(* Logix 5000 project; controller FV vendor 1 type 14 code 217 rev 31.11; software revision 31.00; part 31 of 63 *)
(* tags used below, declared in another part *)
   CWD : CHECKWORD_FLAGS;
   FR_BEACON1 : PlantItem;   // BEACON1
   FR_data_file_value_to_move : DINT;
   FR_F202 : REAL[20];
   FR_F203 : REAL[40];
   FR_N120 : INT[265];   // YEAST CROP Yeast Cropping Main
   FR_N14 : INT[265];   // MVFV CIP Comms to MVFV CIP Un it PLC
   FR_N140 : INT[265];   // CIP
   FR_N160 : INT[265];   // VESSEL Vessel Working Direc tory
   FR_N20 : INT[265];   // GENERAL General Purpose Setp oints
   FR_N30 : INT[265];   // FV30
   FR_N7 : INT[265];   // INTEGER
   FR_N99 : INT[265];   // COMMENT Comment Lines
   FR_T121 : TIMER[255];   // YEAST CROP
   scale_analog_result : REAL;
(* FR_Common, continued *)

ROUTINE FR_VESSEL_160   (* ladder *)
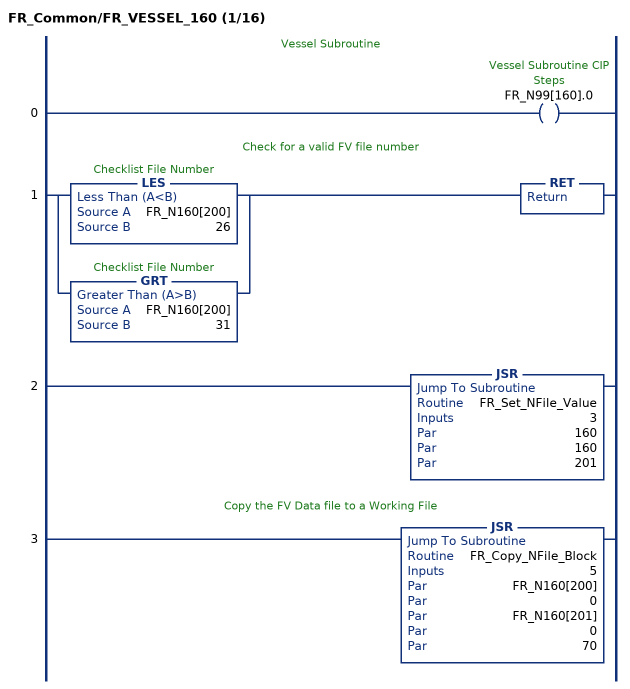
   // Vessel Subroutine
   0: OTE(FR_N99[160].0);
   // Check for a valid FV file number
   1: [LES(FR_N160[200],26) ,GRT(FR_N160[200],31) ]RET();
   2: JSR(FR_Set_NFile_Value,3,160,160,201);
   // Copy the FV Data file to a Working File
   3: JSR(FR_Copy_NFile_Block,5,FR_N160[200],0,FR_N160[201],0,70);
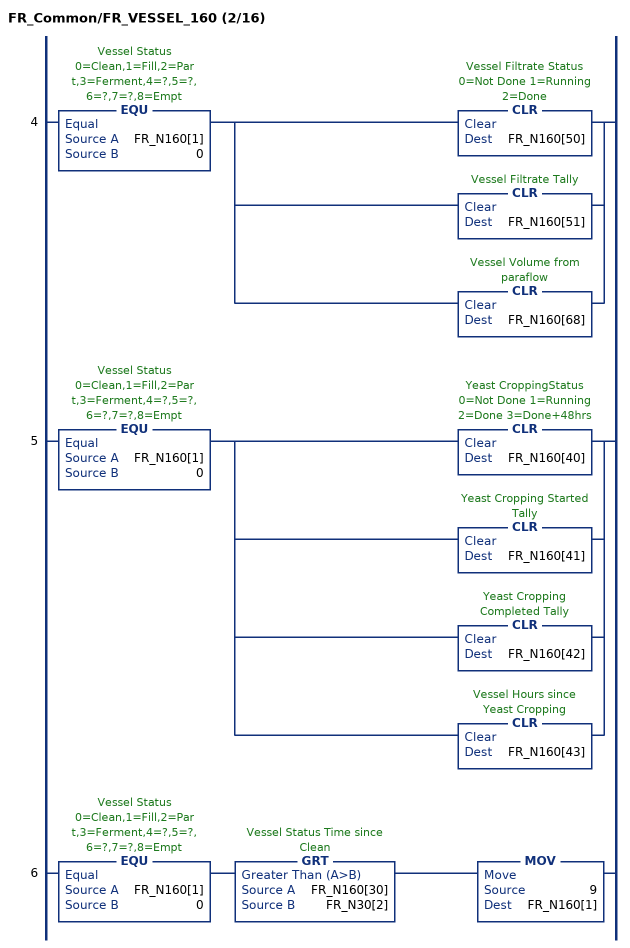
   4: EQU(FR_N160[1],0)[CLR(FR_N160[50]) ,CLR(FR_N160[51]) ,CLR(FR_N160[68]) ];
   5: EQU(FR_N160[1],0)[CLR(FR_N160[40]) ,CLR(FR_N160[41]) ,CLR(FR_N160[42]) ,CLR(FR_N160[43]) ];
   6: EQU(FR_N160[1],0)GRT(FR_N160[30],FR_N30[2])MOV(9,FR_N160[1]);
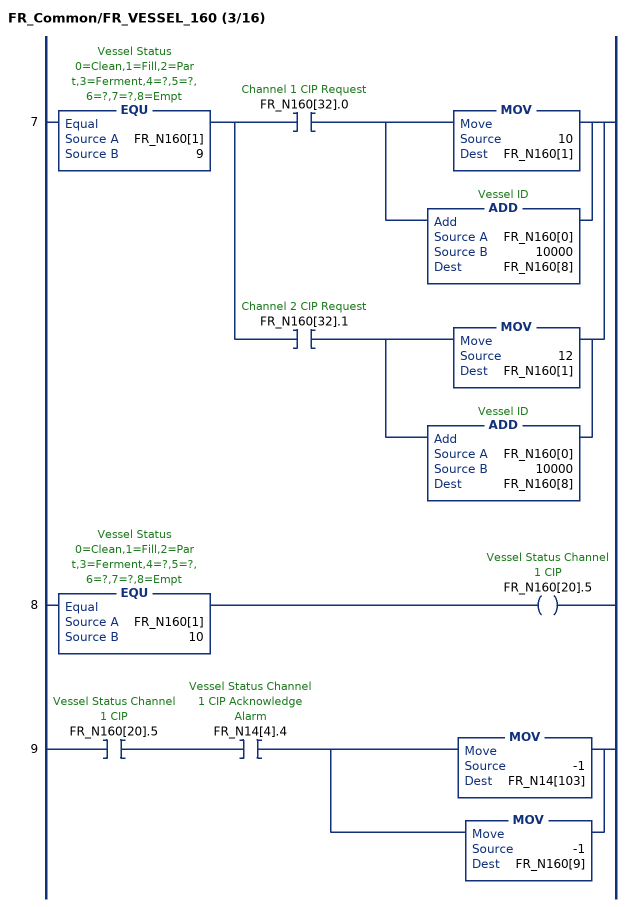
   7: EQU(FR_N160[1],9)[XIC(FR_N160[32].0) [MOV(10,FR_N160[1]) ,ADD(FR_N160[0],10000,FR_N160[8]) ] ,XIC(FR_N160[32].1) [MOV(12,FR_N160[1]) ,ADD(FR_N160[0],10000,FR_N160[8]) ] ];
   8: EQU(FR_N160[1],10)OTE(FR_N160[20].5);
   9: XIC(FR_N160[20].5)XIC(FR_N14[4].4)[MOV(-1,FR_N14[103]) ,MOV(-1,FR_N160[9]) ];
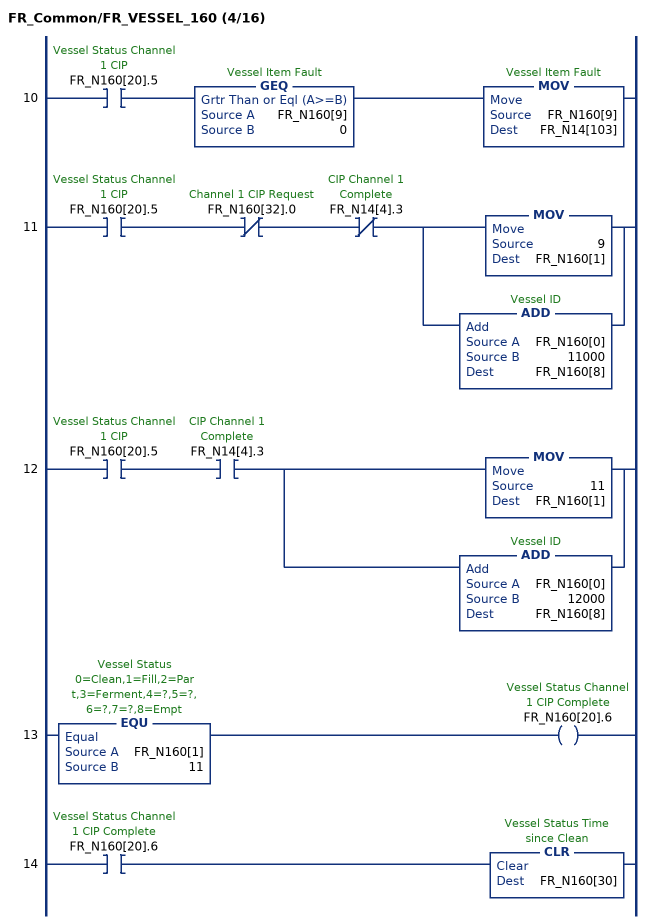
   10: XIC(FR_N160[20].5)GEQ(FR_N160[9],0)MOV(FR_N160[9],FR_N14[103]);
   11: XIC(FR_N160[20].5)XIO(FR_N160[32].0)XIO(FR_N14[4].3)[MOV(9,FR_N160[1]) ,ADD(FR_N160[0],11000,FR_N160[8]) ];
   12: XIC(FR_N160[20].5)XIC(FR_N14[4].3)[MOV(11,FR_N160[1]) ,ADD(FR_N160[0],12000,FR_N160[8]) ];
   13: EQU(FR_N160[1],11)OTE(FR_N160[20].6);
   14: XIC(FR_N160[20].6)CLR(FR_N160[30]);
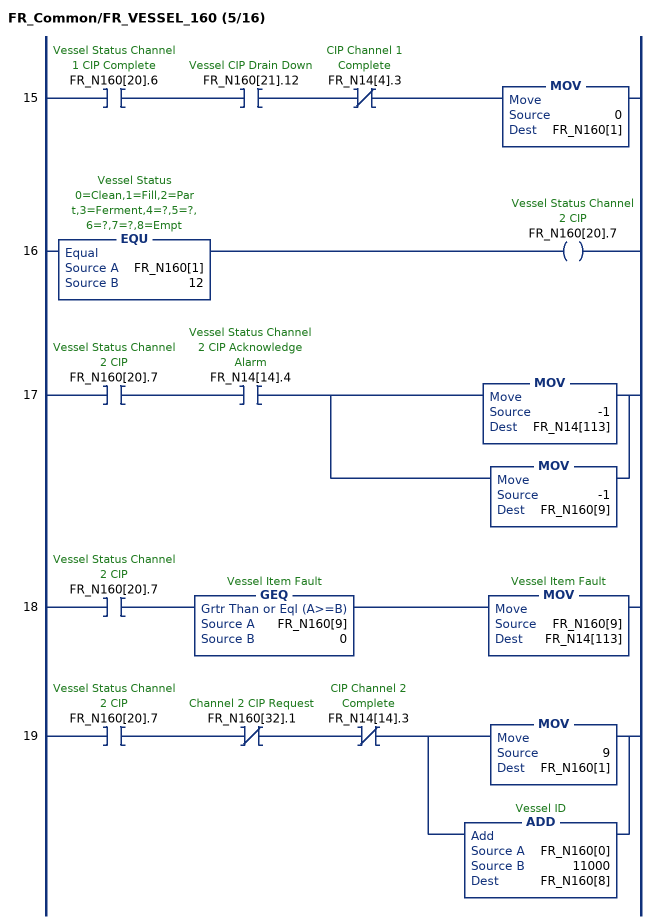
   15: XIC(FR_N160[20].6)XIC(FR_N160[21].12)XIO(FR_N14[4].3)MOV(0,FR_N160[1]);
   16: EQU(FR_N160[1],12)OTE(FR_N160[20].7);
   17: XIC(FR_N160[20].7)XIC(FR_N14[14].4)[MOV(-1,FR_N14[113]) ,MOV(-1,FR_N160[9]) ];
   18: XIC(FR_N160[20].7)GEQ(FR_N160[9],0)MOV(FR_N160[9],FR_N14[113]);
   19: XIC(FR_N160[20].7)XIO(FR_N160[32].1)XIO(FR_N14[14].3)[MOV(9,FR_N160[1]) ,ADD(FR_N160[0],11000,FR_N160[8]) ];
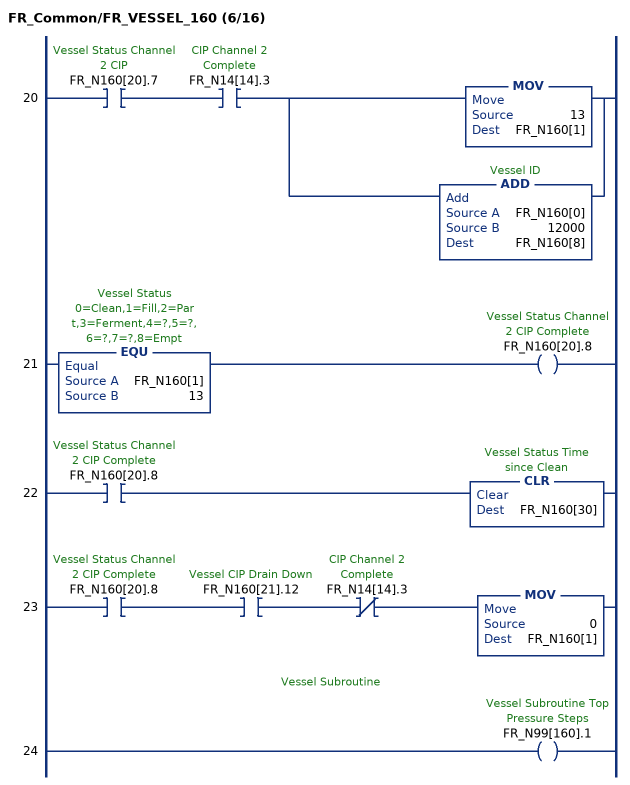
   20: XIC(FR_N160[20].7)XIC(FR_N14[14].3)[MOV(13,FR_N160[1]) ,ADD(FR_N160[0],12000,FR_N160[8]) ];
   21: EQU(FR_N160[1],13)OTE(FR_N160[20].8);
   22: XIC(FR_N160[20].8)CLR(FR_N160[30]);
   23: XIC(FR_N160[20].8)XIC(FR_N160[21].12)XIO(FR_N14[14].3)MOV(0,FR_N160[1]);
   // Vessel Subroutine
   24: OTE(FR_N99[160].1);
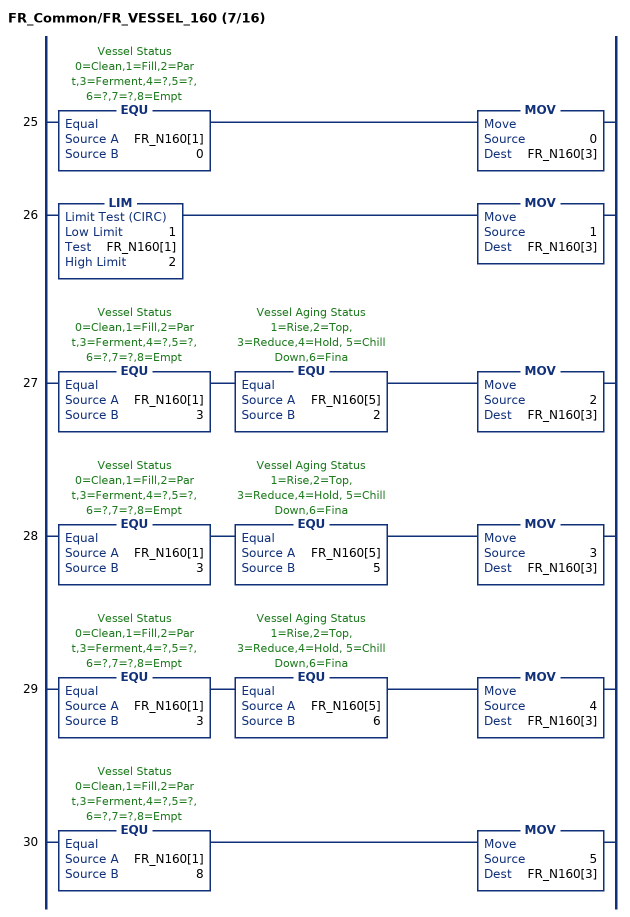
   25: EQU(FR_N160[1],0)MOV(0,FR_N160[3]);
   26: LIM(1,FR_N160[1],2)MOV(1,FR_N160[3]);
   27: EQU(FR_N160[1],3)EQU(FR_N160[5],2)MOV(2,FR_N160[3]);
   28: EQU(FR_N160[1],3)EQU(FR_N160[5],5)MOV(3,FR_N160[3]);
   29: EQU(FR_N160[1],3)EQU(FR_N160[5],6)MOV(4,FR_N160[3]);
   30: EQU(FR_N160[1],8)MOV(5,FR_N160[3]);
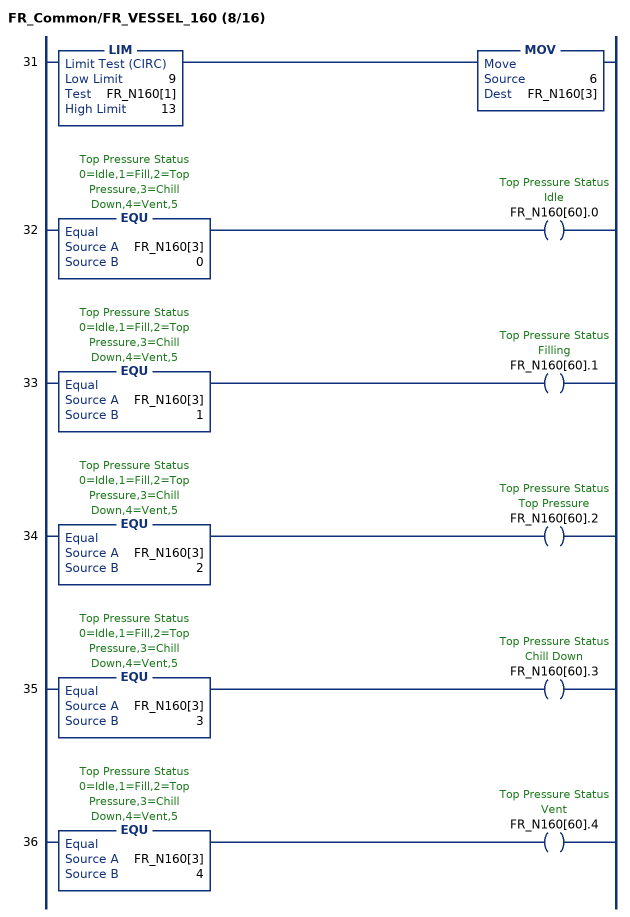
   31: LIM(9,FR_N160[1],13)MOV(6,FR_N160[3]);
   32: EQU(FR_N160[3],0)OTE(FR_N160[60].0);
   33: EQU(FR_N160[3],1)OTE(FR_N160[60].1);
   34: EQU(FR_N160[3],2)OTE(FR_N160[60].2);
   35: EQU(FR_N160[3],3)OTE(FR_N160[60].3);
   36: EQU(FR_N160[3],4)OTE(FR_N160[60].4);
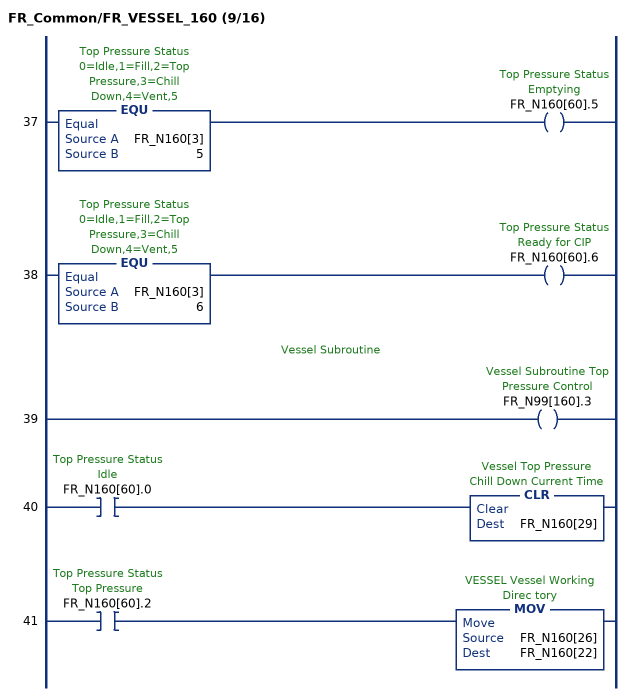
   37: EQU(FR_N160[3],5)OTE(FR_N160[60].5);
   38: EQU(FR_N160[3],6)OTE(FR_N160[60].6);
   // Vessel Subroutine
   39: OTE(FR_N99[160].3);
   40: XIC(FR_N160[60].0)CLR(FR_N160[29]);
   41: XIC(FR_N160[60].2)MOV(FR_N160[26],FR_N160[22]);
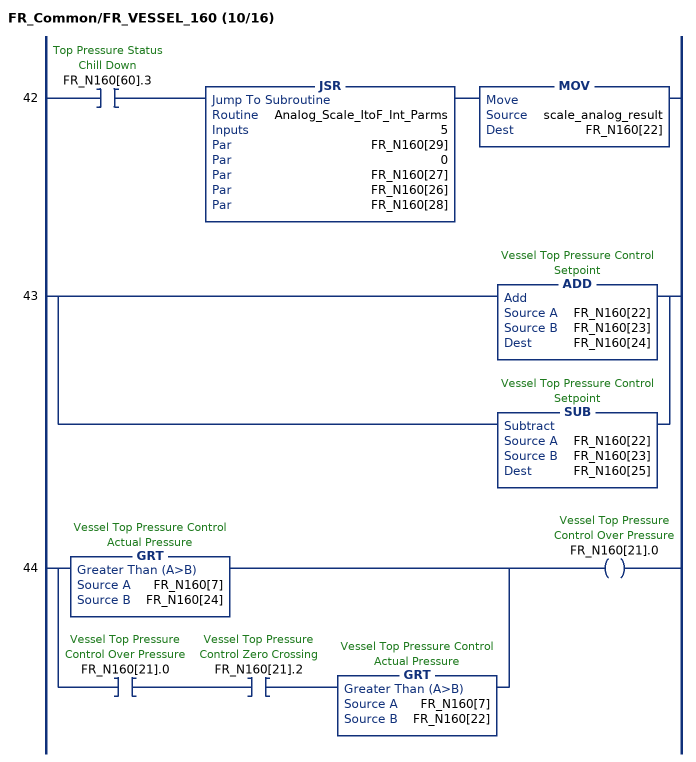
   42: XIC(FR_N160[60].3)JSR(Analog_Scale_ItoF_Int_Parms,5,FR_N160[29],0,FR_N160[27],FR_N160[26],FR_N160[28])MOV(scale_analog_result,FR_N160[22]);
   43: [ADD(FR_N160[22],FR_N160[23],FR_N160[24]) ,SUB(FR_N160[22],FR_N160[23],FR_N160[25]) ];
   44: [GRT(FR_N160[7],FR_N160[24]) ,XIC(FR_N160[21].0) XIC(FR_N160[21].2) GRT(FR_N160[7],FR_N160[22]) ]OTE(FR_N160[21].0);
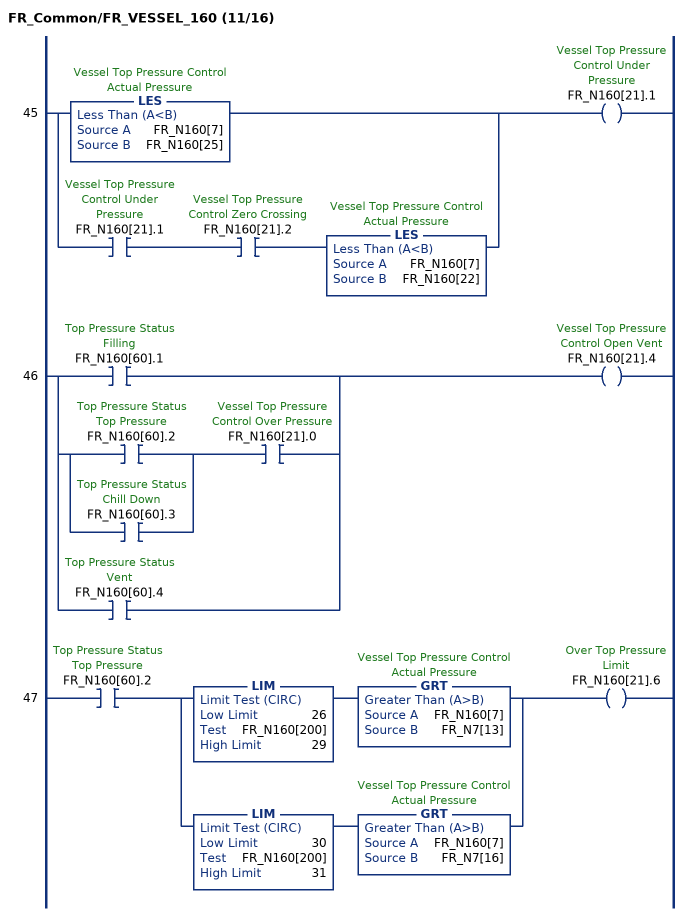
   45: [LES(FR_N160[7],FR_N160[25]) ,XIC(FR_N160[21].1) XIC(FR_N160[21].2) LES(FR_N160[7],FR_N160[22]) ]OTE(FR_N160[21].1);
   46: [XIC(FR_N160[60].1) ,[XIC(FR_N160[60].2) ,XIC(FR_N160[60].3) ] XIC(FR_N160[21].0) ,XIC(FR_N160[60].4) ]OTE(FR_N160[21].4);
   47: XIC(FR_N160[60].2)[LIM(26,FR_N160[200],29) GRT(FR_N160[7],FR_N7[13]) ,LIM(30,FR_N160[200],31) GRT(FR_N160[7],FR_N7[16]) ]OTE(FR_N160[21].6);
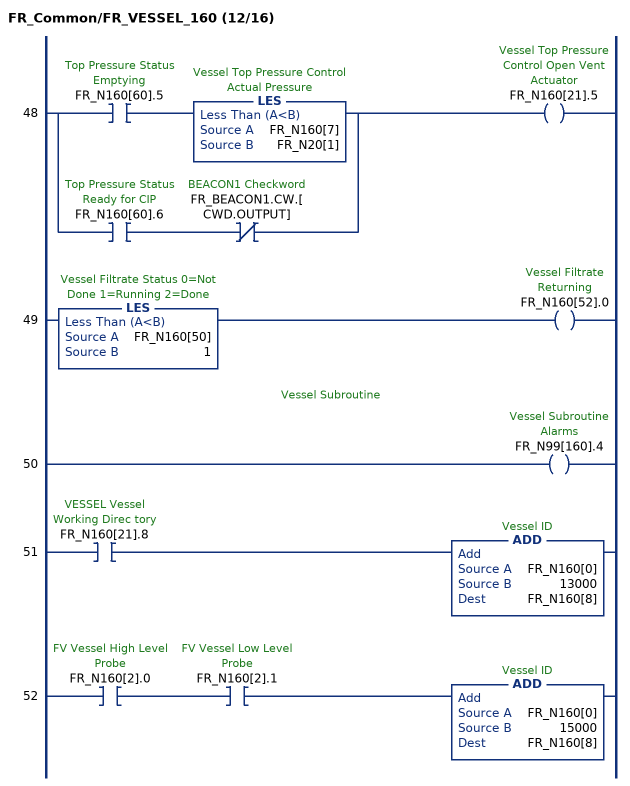
   48: [XIC(FR_N160[60].5) LES(FR_N160[7],FR_N20[1]) ,XIC(FR_N160[60].6) XIO(FR_BEACON1.CW.[CWD.OUTPUT]) ]OTE(FR_N160[21].5);
   49: LES(FR_N160[50],1)OTE(FR_N160[52].0);
   // Vessel Subroutine
   50: OTE(FR_N99[160].4);
   51: XIC(FR_N160[21].8)ADD(FR_N160[0],13000,FR_N160[8]);
   52: XIC(FR_N160[2].0)XIC(FR_N160[2].1)ADD(FR_N160[0],15000,FR_N160[8]);
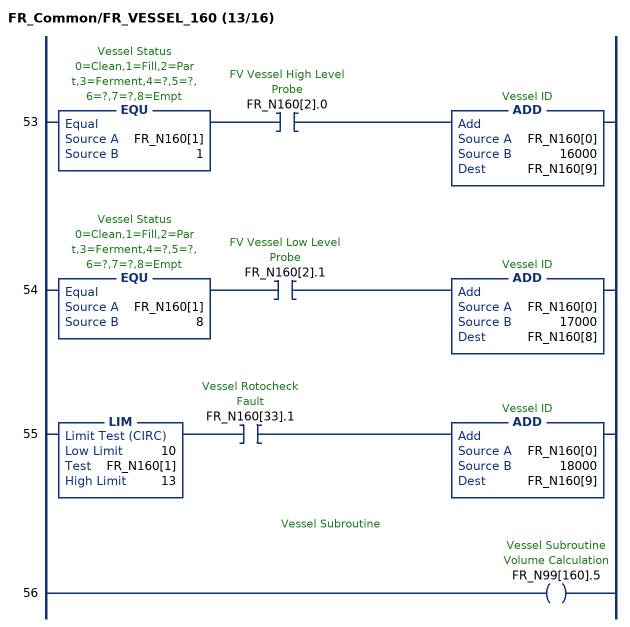
   53: EQU(FR_N160[1],1)XIC(FR_N160[2].0)ADD(FR_N160[0],16000,FR_N160[9]);
   54: EQU(FR_N160[1],8)XIC(FR_N160[2].1)ADD(FR_N160[0],17000,FR_N160[8]);
   55: LIM(10,FR_N160[1],13)XIC(FR_N160[33].1)ADD(FR_N160[0],18000,FR_N160[9]);
   // Vessel Subroutine
   56: OTE(FR_N99[160].5);
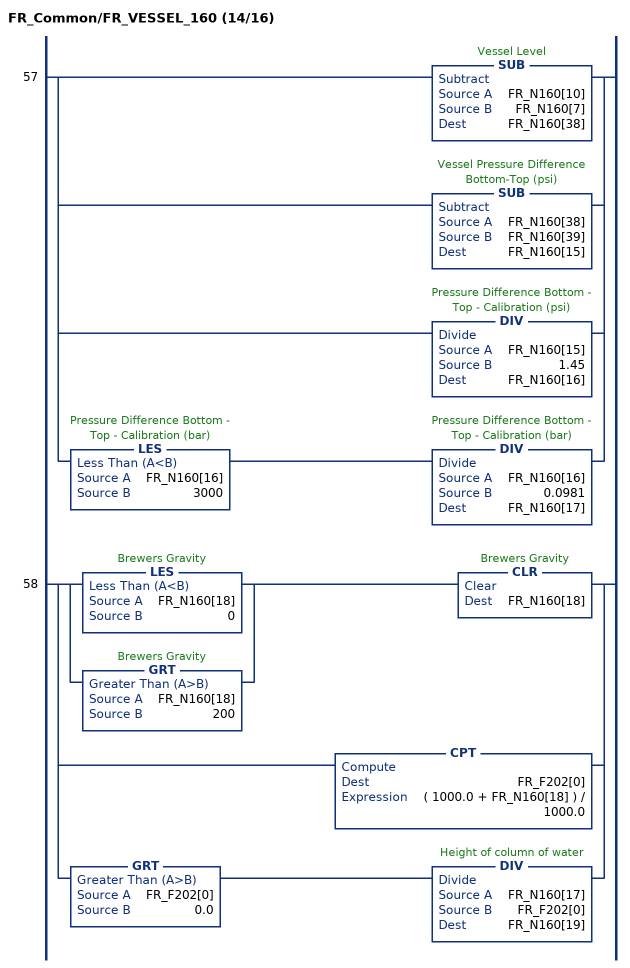
   57: [SUB(FR_N160[10],FR_N160[7],FR_N160[38]) ,SUB(FR_N160[38],FR_N160[39],FR_N160[15]) ,DIV(FR_N160[15],1.45,FR_N160[16]) ,LES(FR_N160[16],3000) DIV(FR_N160[16],0.0981,FR_N160[17]) ];
   58: [[LES(FR_N160[18],0) ,GRT(FR_N160[18],200) ] CLR(FR_N160[18]) ,CPT(FR_F202[0],( 1000.0 + FR_N160[18] ) / 1000.0) ,GRT(FR_F202[0],0.0) DIV(FR_N160[17],FR_F202[0],FR_N160[19]) ];
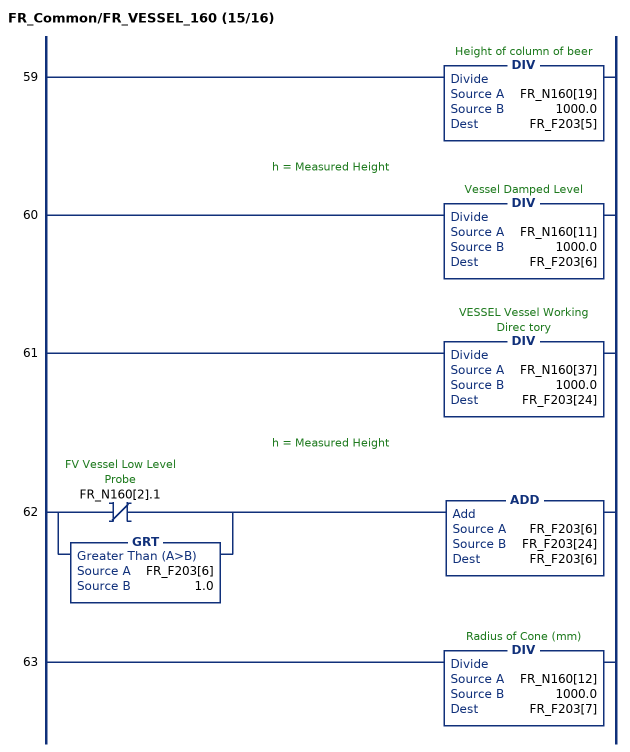
   59: DIV(FR_N160[19],1000.0,FR_F203[5]);
   // h = Measured Height
   60: DIV(FR_N160[11],1000.0,FR_F203[6]);
   61: DIV(FR_N160[37],1000.0,FR_F203[24]);
   // h = Measured Height
   62: [XIO(FR_N160[2].1) ,GRT(FR_F203[6],1.0) ]ADD(FR_F203[6],FR_F203[24],FR_F203[6]);
   63: DIV(FR_N160[12],1000.0,FR_F203[7]);
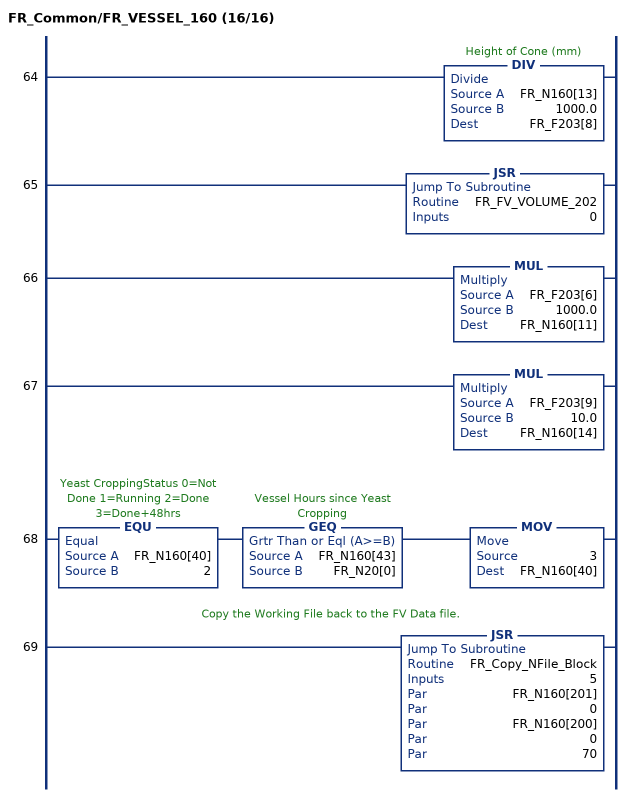
   64: DIV(FR_N160[13],1000.0,FR_F203[8]);
   65: JSR(FR_FV_VOLUME_202,0);
   66: MUL(FR_F203[6],1000.0,FR_N160[11]);
   67: MUL(FR_F203[9],10.0,FR_N160[14]);
   68: EQU(FR_N160[40],2)GEQ(FR_N160[43],FR_N20[0])MOV(3,FR_N160[40]);
   // Copy the Working File back to the FV Data file.
   69: JSR(FR_Copy_NFile_Block,5,FR_N160[201],0,FR_N160[200],0,70);
END_ROUTINE

ROUTINE FR_YEAST_121   (* ladder *)
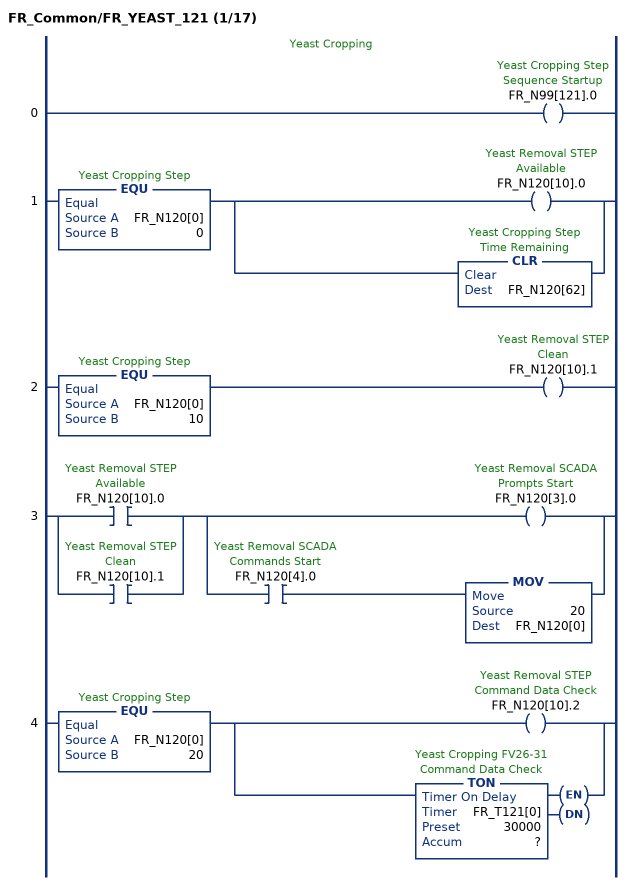
   // Yeast Cropping
   0: OTE(FR_N99[121].0);
   1: EQU(FR_N120[0],0)[OTE(FR_N120[10].0) ,CLR(FR_N120[62]) ];
   2: EQU(FR_N120[0],10)OTE(FR_N120[10].1);
   3: [XIC(FR_N120[10].0) ,XIC(FR_N120[10].1) ][OTE(FR_N120[3].0) ,XIC(FR_N120[4].0) MOV(20,FR_N120[0]) ];
   4: EQU(FR_N120[0],20)[OTE(FR_N120[10].2) ,TON(FR_T121[0],?,?) ];
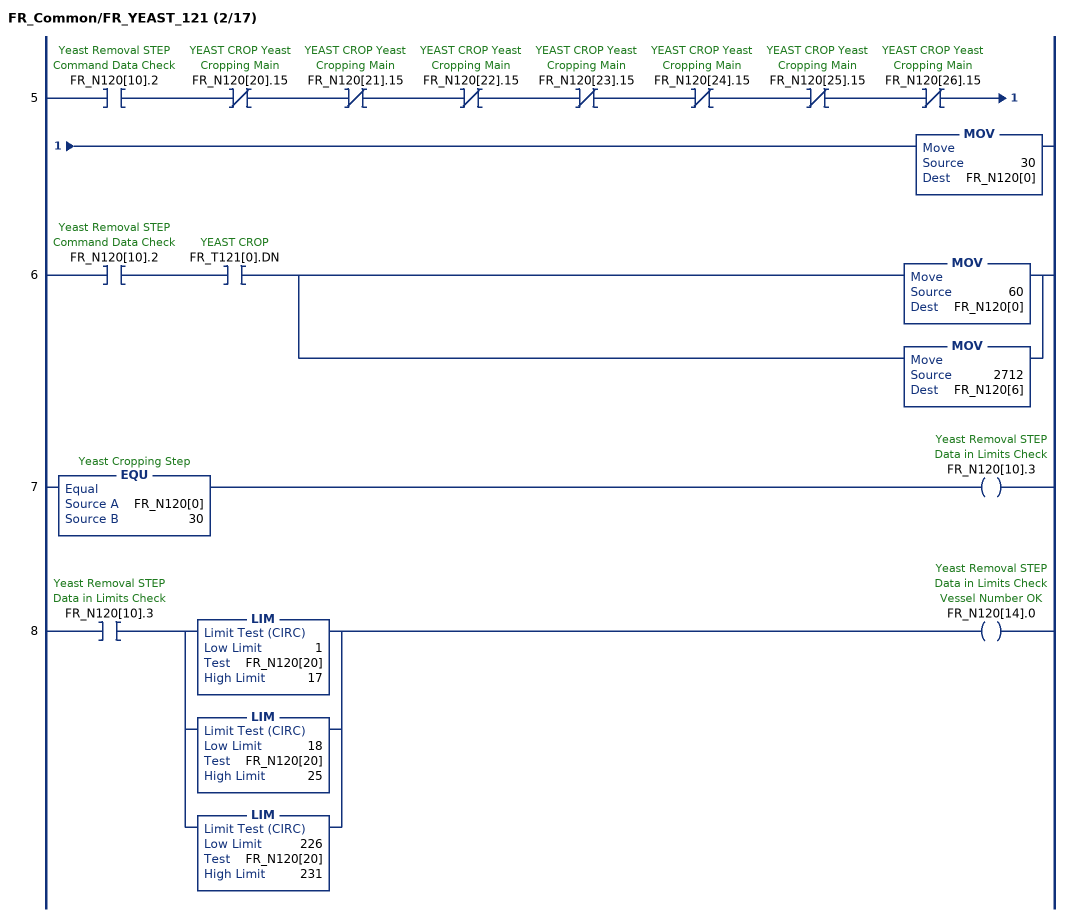
   5: XIC(FR_N120[10].2)XIO(FR_N120[20].15)XIO(FR_N120[21].15)XIO(FR_N120[22].15)XIO(FR_N120[23].15)XIO(FR_N120[24].15)XIO(FR_N120[25].15)XIO(FR_N120[26].15)MOV(30,FR_N120[0]);
   6: XIC(FR_N120[10].2)XIC(FR_T121[0].DN)[MOV(60,FR_N120[0]) ,MOV(2712,FR_N120[6]) ];
   7: EQU(FR_N120[0],30)OTE(FR_N120[10].3);
   8: XIC(FR_N120[10].3)[LIM(1,FR_N120[20],17) ,LIM(18,FR_N120[20],25) ,LIM(226,FR_N120[20],231) ]OTE(FR_N120[14].0);
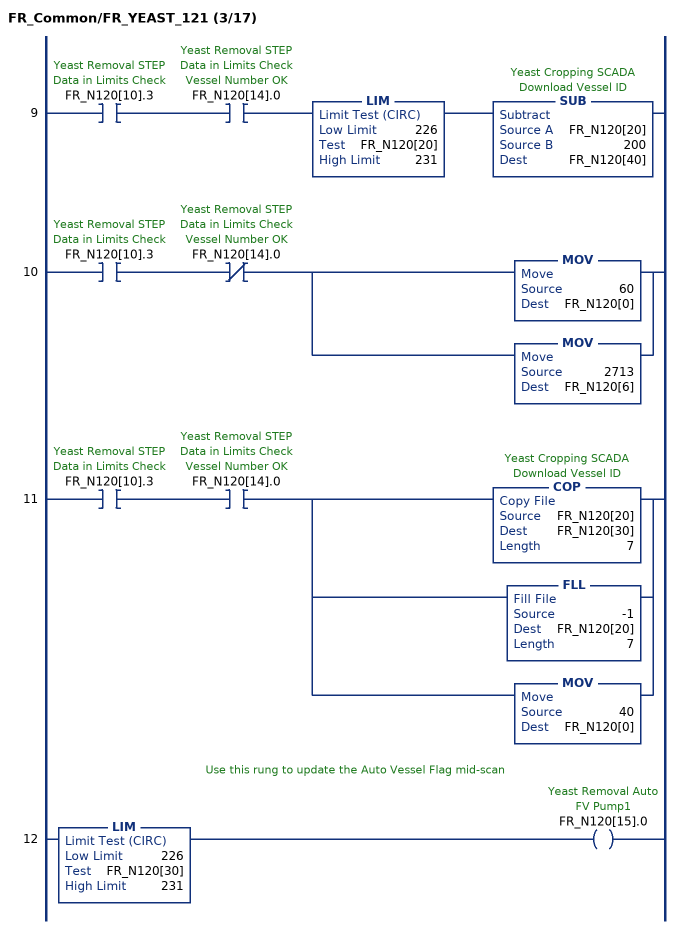
   9: XIC(FR_N120[10].3)XIC(FR_N120[14].0)LIM(226,FR_N120[20],231)SUB(FR_N120[20],200,FR_N120[40]);
   10: XIC(FR_N120[10].3)XIO(FR_N120[14].0)[MOV(60,FR_N120[0]) ,MOV(2713,FR_N120[6]) ];
   11: XIC(FR_N120[10].3)XIC(FR_N120[14].0)[COP(FR_N120[20],FR_N120[30],7) ,FLL(-1,FR_N120[20],7) ,MOV(40,FR_N120[0]) ];
   // Use this rung to update the Auto Vessel Flag mid-scan
   12: LIM(226,FR_N120[30],231)OTE(FR_N120[15].0);
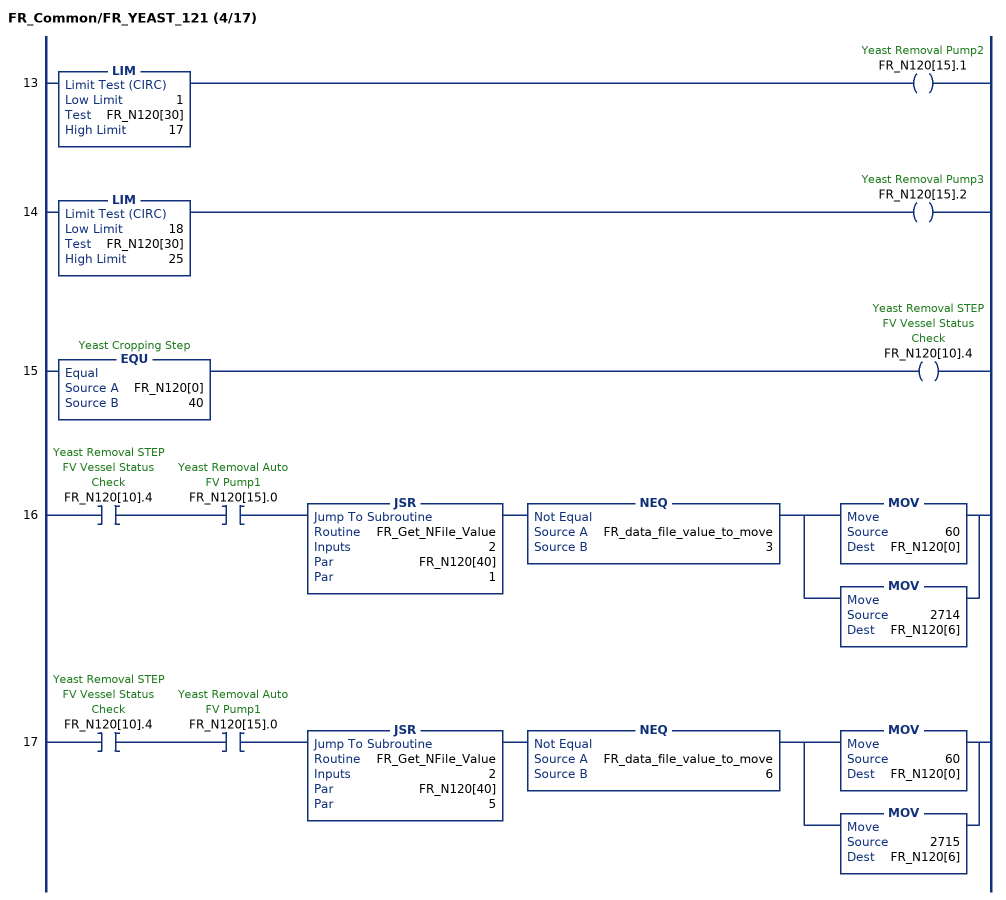
   13: LIM(1,FR_N120[30],17)OTE(FR_N120[15].1);
   14: LIM(18,FR_N120[30],25)OTE(FR_N120[15].2);
   15: EQU(FR_N120[0],40)OTE(FR_N120[10].4);
   16: XIC(FR_N120[10].4)XIC(FR_N120[15].0)JSR(FR_Get_NFile_Value,2,FR_N120[40],1)NEQ(FR_data_file_value_to_move,3)[MOV(60,FR_N120[0]) ,MOV(2714,FR_N120[6]) ];
   17: XIC(FR_N120[10].4)XIC(FR_N120[15].0)JSR(FR_Get_NFile_Value,2,FR_N120[40],5)NEQ(FR_data_file_value_to_move,6)[MOV(60,FR_N120[0]) ,MOV(2715,FR_N120[6]) ];
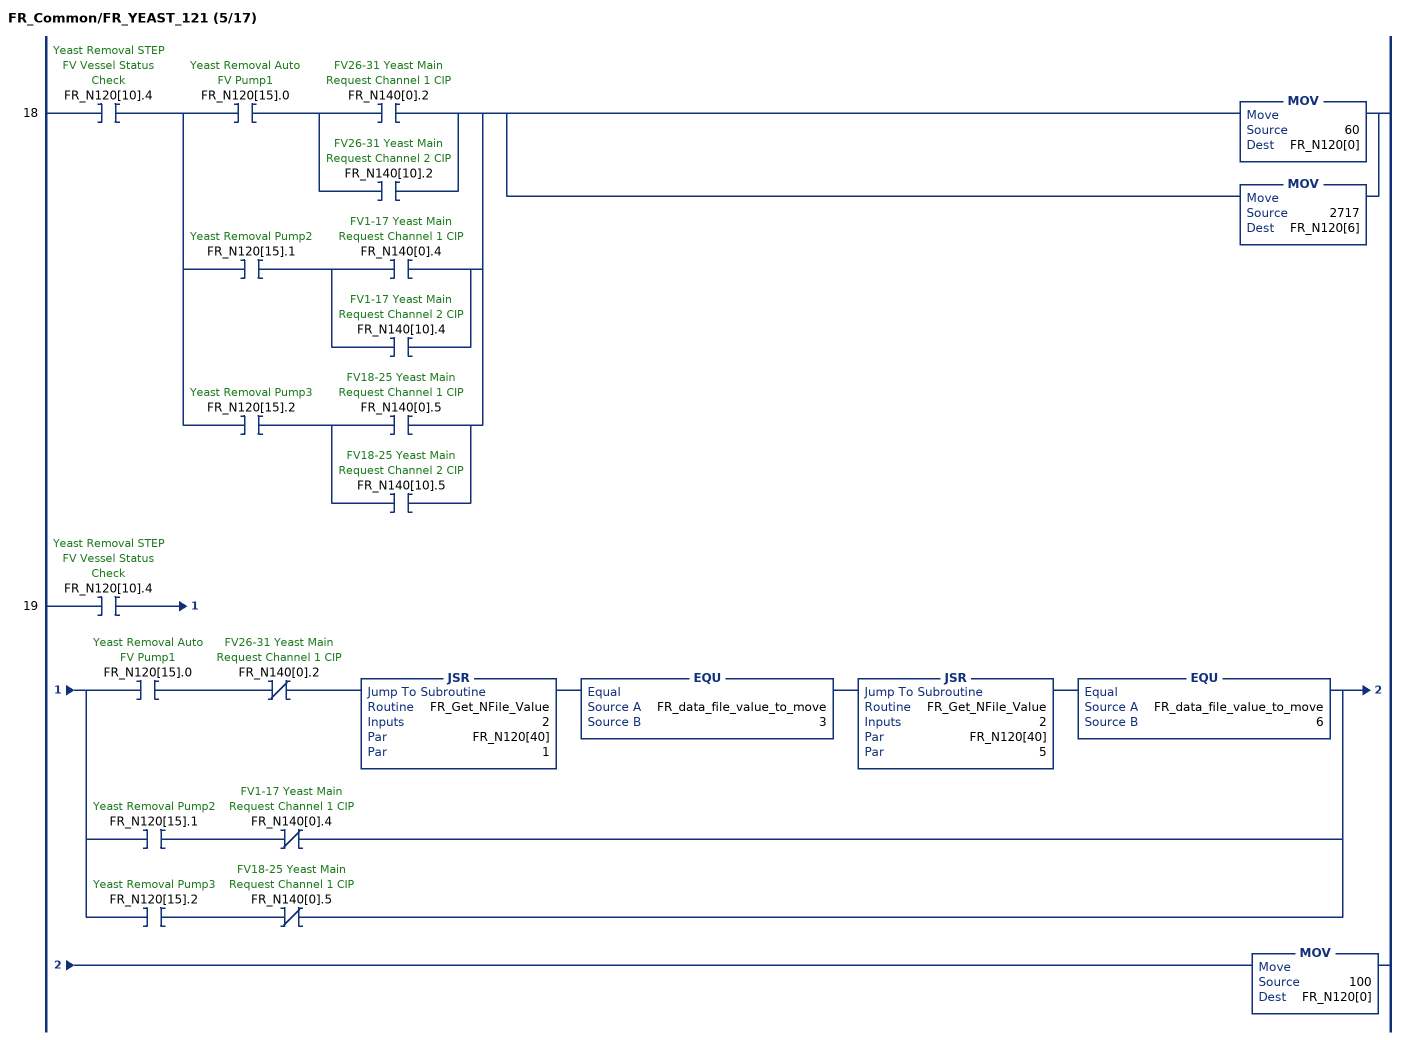
   18: XIC(FR_N120[10].4)[XIC(FR_N120[15].0) [XIC(FR_N140[0].2) ,XIC(FR_N140[10].2) ] ,XIC(FR_N120[15].1) [XIC(FR_N140[0].4) ,XIC(FR_N140[10].4) ] ,XIC(FR_N120[15].2) [XIC(FR_N140[0].5) ,XIC(FR_N140[10].5) ] ][MOV(60,FR_N120[0]) ,MOV(2717,FR_N120[6]) ];
   19: XIC(FR_N120[10].4)[XIC(FR_N120[15].0) XIO(FR_N140[0].2) JSR(FR_Get_NFile_Value,2,FR_N120[40],1) EQU(FR_data_file_value_to_move,3) JSR(FR_Get_NFile_Value,2,FR_N120[40],5) EQU(FR_data_file_value_to_move,6) ,XIC(FR_N120[15].1) XIO(FR_N140[0].4) ,XIC(FR_N120[15].2) XIO(FR_N140[0].5) ]MOV(100,FR_N120[0]);
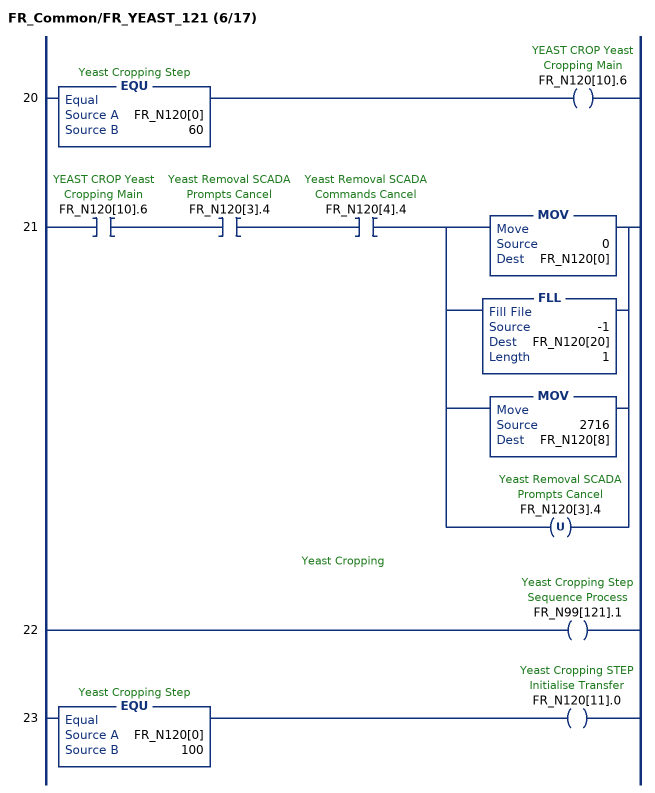
   20: EQU(FR_N120[0],60)OTE(FR_N120[10].6);
   21: XIC(FR_N120[10].6)XIC(FR_N120[3].4)XIC(FR_N120[4].4)[MOV(0,FR_N120[0]) ,FLL(-1,FR_N120[20],1) ,MOV(2716,FR_N120[8]) ,OTU(FR_N120[3].4) ];
   // Yeast Cropping
   22: OTE(FR_N99[121].1);
   23: EQU(FR_N120[0],100)OTE(FR_N120[11].0);
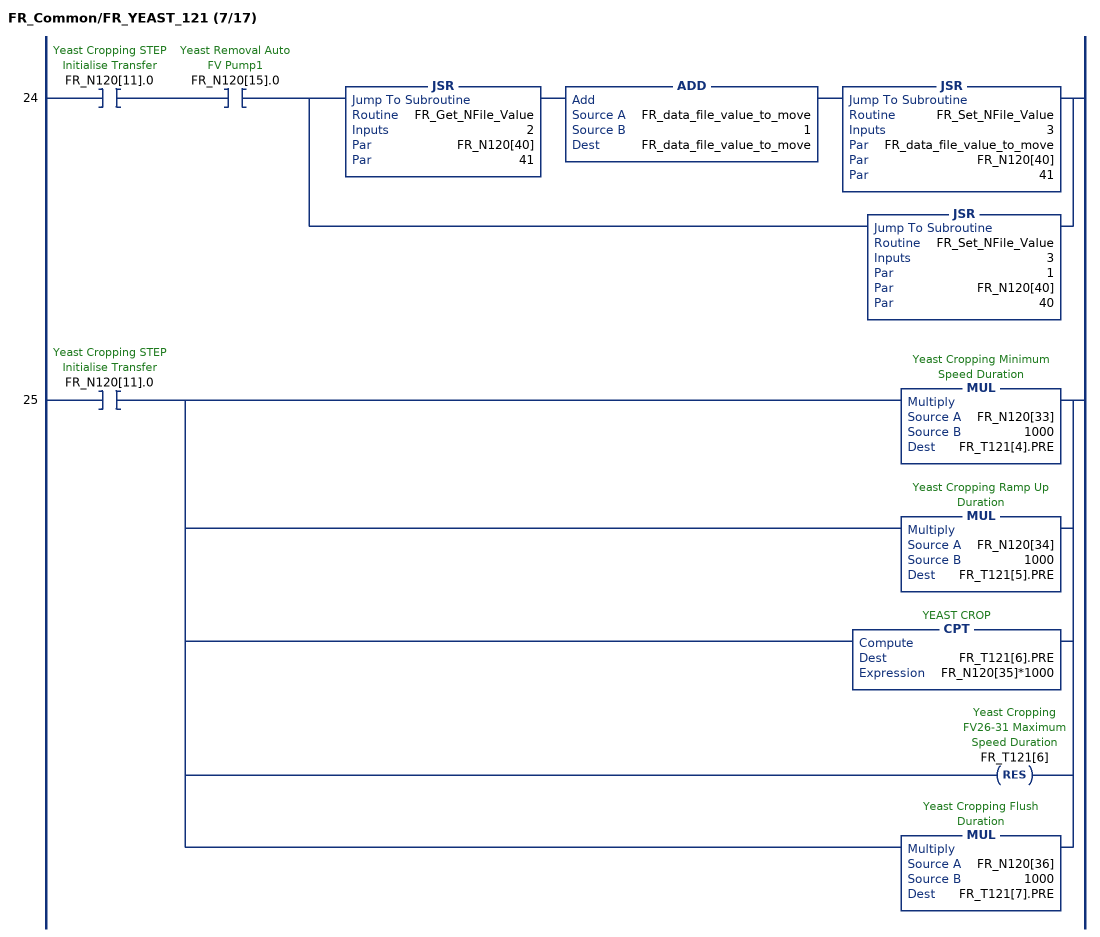
   24: XIC(FR_N120[11].0)XIC(FR_N120[15].0)[JSR(FR_Get_NFile_Value,2,FR_N120[40],41) ADD(FR_data_file_value_to_move,1,FR_data_file_value_to_move) JSR(FR_Set_NFile_Value,3,FR_data_file_value_to_move,FR_N120[40],41) ,JSR(FR_Set_NFile_Value,3,1,FR_N120[40],40) ];
   25: XIC(FR_N120[11].0)[MUL(FR_N120[33],1000,FR_T121[4].PRE) ,MUL(FR_N120[34],1000,FR_T121[5].PRE) ,CPT(FR_T121[6].PRE,FR_N120[35]*1000) ,RES(FR_T121[6]) ,MUL(FR_N120[36],1000,FR_T121[7].PRE) ];
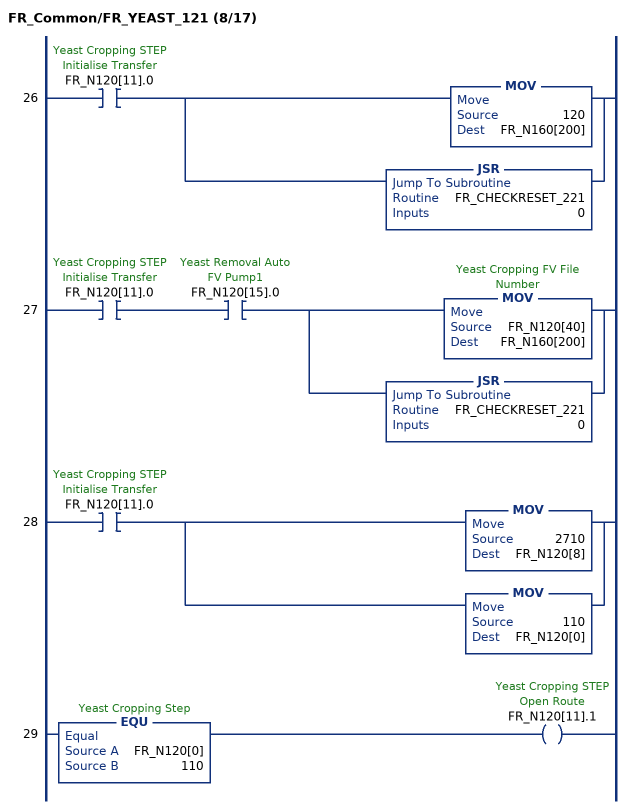
   26: XIC(FR_N120[11].0)[MOV(120,FR_N160[200]) ,JSR(FR_CHECKRESET_221,0) ];
   27: XIC(FR_N120[11].0)XIC(FR_N120[15].0)[MOV(FR_N120[40],FR_N160[200]) ,JSR(FR_CHECKRESET_221,0) ];
   28: XIC(FR_N120[11].0)[MOV(2710,FR_N120[8]) ,MOV(110,FR_N120[0]) ];
   29: EQU(FR_N120[0],110)OTE(FR_N120[11].1);
